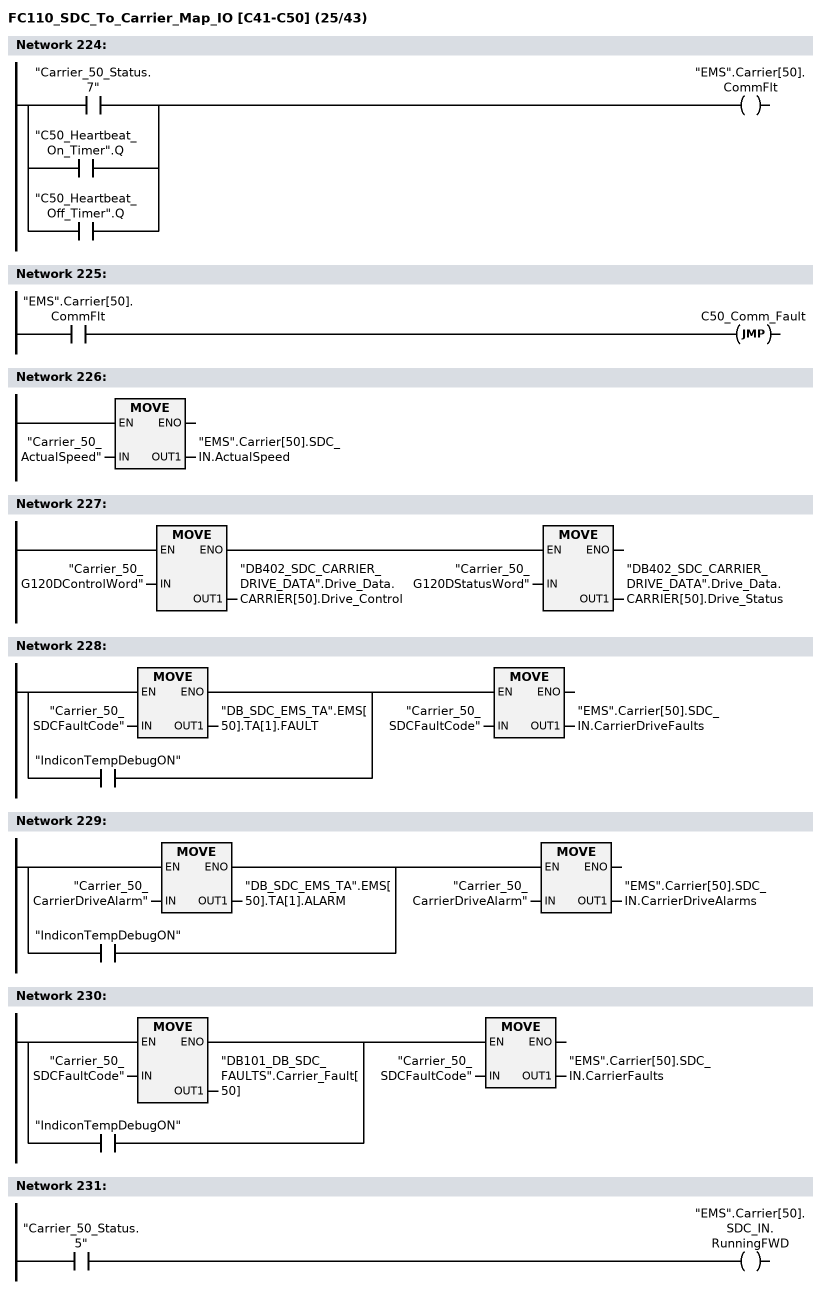
   RUNG wire#powerrail
      Contact( "Carrier_50_Status.7" )
      wire#w1
      Coil( "EMS".Carrier[50].CommFlt )
   END_RUNG
   RUNG wire#powerrail
      Contact( "C50_Heartbeat_On_Timer".Q )
   END_RUNG wire#w1
   RUNG wire#powerrail
      Contact( "C50_Heartbeat_Off_Timer".Q )
   END_RUNG wire#w1
   // the same network as SCL:
   "EMS".Carrier[50].CommFlt := "Carrier_50_Status.7" OR "C50_Heartbeat_On_Timer".Q OR "C50_Heartbeat_Off_Timer".Q;
END_REGION

REGION Network 225
   RUNG wire#powerrail
      Contact( "EMS".Carrier[50].CommFlt )
      JumpCoil( C50_Comm_Fault )
   END_RUNG
   // the same network as SCL:
   IF "EMS".Carrier[50].CommFlt THEN GOTO C50_Comm_Fault; END_IF;
END_REGION

REGION Network 226
   RUNG wire#powerrail
      Move(in := "Carrier_50_ActualSpeed", out1 => "EMS".Carrier[50].SDC_IN.ActualSpeed)
   END_RUNG
   // the same network as SCL:
   "EMS".Carrier[50].SDC_IN.ActualSpeed := "Carrier_50_ActualSpeed";
END_REGION

REGION Network 227
   RUNG wire#powerrail
      Move(in := "Carrier_50_G120DControlWord", out1 => "DB402_SDC_CARRIER_DRIVE_DATA".Drive_Data.CARRIER[50].Drive_Control)
      Move(in := "Carrier_50_G120DStatusWord", out1 => "DB402_SDC_CARRIER_DRIVE_DATA".Drive_Data.CARRIER[50].Drive_Status)
   END_RUNG
   // the same network as SCL:
   "DB402_SDC_CARRIER_DRIVE_DATA".Drive_Data.CARRIER[50].Drive_Control := "Carrier_50_G120DControlWord";
   "DB402_SDC_CARRIER_DRIVE_DATA".Drive_Data.CARRIER[50].Drive_Status := "Carrier_50_G120DStatusWord";
END_REGION

REGION Network 228
   RUNG wire#powerrail
      Move(in := "Carrier_50_SDCFaultCode", out1 => "DB_SDC_EMS_TA".EMS[50].TA[1].FAULT)
      wire#w1
      Move(in := "Carrier_50_SDCFaultCode", out1 => "EMS".Carrier[50].SDC_IN.CarrierDriveFaults)
   END_RUNG
   RUNG wire#powerrail
      Contact( "IndiconTempDebugON" )
   END_RUNG wire#w1
   // the same network as SCL:
   "DB_SDC_EMS_TA".EMS[50].TA[1].FAULT := "Carrier_50_SDCFaultCode";
   IF TRUE OR "IndiconTempDebugON" THEN
       "EMS".Carrier[50].SDC_IN.CarrierDriveFaults := "Carrier_50_SDCFaultCode";
   END_IF;
END_REGION

REGION Network 229
   RUNG wire#powerrail
      Move(in := "Carrier_50_CarrierDriveAlarm", out1 => "DB_SDC_EMS_TA".EMS[50].TA[1].ALARM)
      wire#w1
      Move(in := "Carrier_50_CarrierDriveAlarm", out1 => "EMS".Carrier[50].SDC_IN.CarrierDriveAlarms)
   END_RUNG
   RUNG wire#powerrail
      Contact( "IndiconTempDebugON" )
   END_RUNG wire#w1
   // the same network as SCL:
   "DB_SDC_EMS_TA".EMS[50].TA[1].ALARM := "Carrier_50_CarrierDriveAlarm";
   IF TRUE OR "IndiconTempDebugON" THEN
       "EMS".Carrier[50].SDC_IN.CarrierDriveAlarms := "Carrier_50_CarrierDriveAlarm";
   END_IF;
END_REGION

REGION Network 230
   RUNG wire#powerrail
      Move(in := "Carrier_50_SDCFaultCode", out1 => "DB101_DB_SDC_FAULTS".Carrier_Fault[50])
      wire#w1
      Move(in := "Carrier_50_SDCFaultCode", out1 => "EMS".Carrier[50].SDC_IN.CarrierFaults)
   END_RUNG
   RUNG wire#powerrail
      Contact( "IndiconTempDebugON" )
   END_RUNG wire#w1
   // the same network as SCL:
   "DB101_DB_SDC_FAULTS".Carrier_Fault[50] := "Carrier_50_SDCFaultCode";
   IF TRUE OR "IndiconTempDebugON" THEN
       "EMS".Carrier[50].SDC_IN.CarrierFaults := "Carrier_50_SDCFaultCode";
   END_IF;
END_REGION

REGION Network 231
   RUNG wire#powerrail
      Contact( "Carrier_50_Status.5" )
      Coil( "EMS".Carrier[50].SDC_IN.RunningFWD )
   END_RUNG
   // the same network as SCL:
   "EMS".Carrier[50].SDC_IN.RunningFWD := "Carrier_50_Status.5";
END_REGION

REGION Network 232
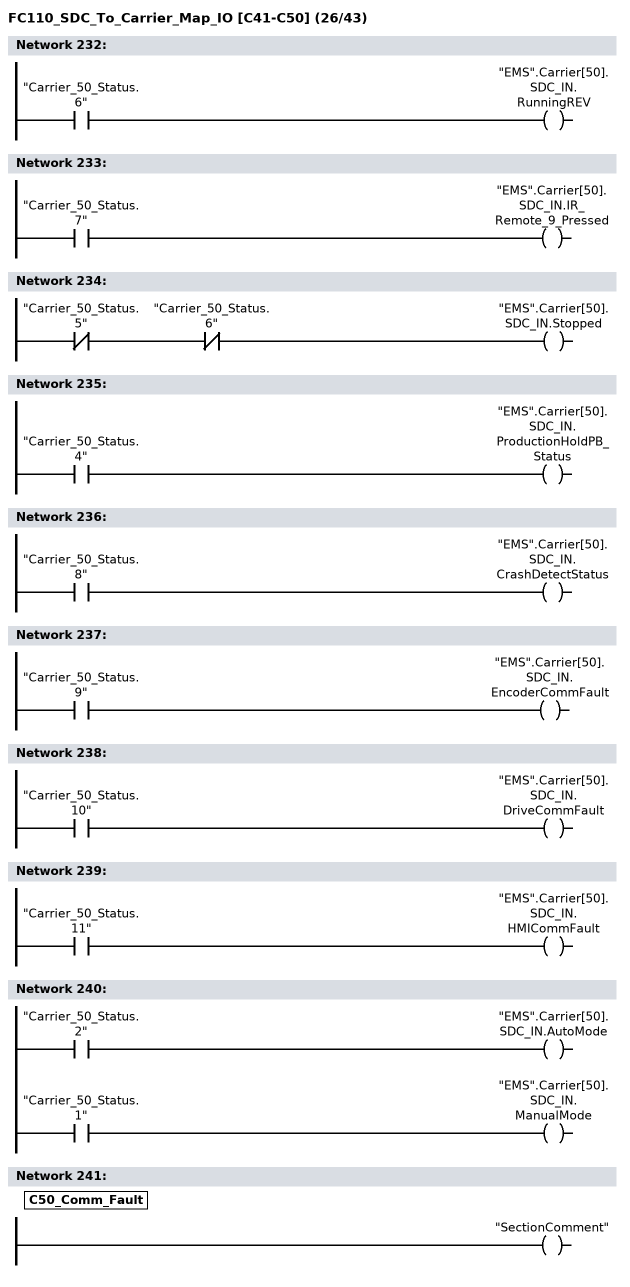
   RUNG wire#powerrail
      Contact( "Carrier_50_Status.6" )
      Coil( "EMS".Carrier[50].SDC_IN.RunningREV )
   END_RUNG
   // the same network as SCL:
   "EMS".Carrier[50].SDC_IN.RunningREV := "Carrier_50_Status.6";
END_REGION

REGION Network 233
   RUNG wire#powerrail
      Contact( "Carrier_50_Status.7" )
      Coil( "EMS".Carrier[50].SDC_IN.IR_Remote_9_Pressed )
   END_RUNG
   // the same network as SCL:
   "EMS".Carrier[50].SDC_IN.IR_Remote_9_Pressed := "Carrier_50_Status.7";
END_REGION

REGION Network 234
   RUNG wire#powerrail
      I_Contact( "Carrier_50_Status.5" )
      I_Contact( "Carrier_50_Status.6" )
      Coil( "EMS".Carrier[50].SDC_IN.Stopped )
   END_RUNG
   // the same network as SCL:
   "EMS".Carrier[50].SDC_IN.Stopped := NOT "Carrier_50_Status.5" AND NOT "Carrier_50_Status.6";
END_REGION

REGION Network 235
   RUNG wire#powerrail
      Contact( "Carrier_50_Status.4" )
      Coil( "EMS".Carrier[50].SDC_IN.ProductionHoldPB_Status )
   END_RUNG
   // the same network as SCL:
   "EMS".Carrier[50].SDC_IN.ProductionHoldPB_Status := "Carrier_50_Status.4";
END_REGION

REGION Network 236
   RUNG wire#powerrail
      Contact( "Carrier_50_Status.8" )
      Coil( "EMS".Carrier[50].SDC_IN.CrashDetectStatus )
   END_RUNG
   // the same network as SCL:
   "EMS".Carrier[50].SDC_IN.CrashDetectStatus := "Carrier_50_Status.8";
END_REGION

REGION Network 237
   RUNG wire#powerrail
      Contact( "Carrier_50_Status.9" )
      Coil( "EMS".Carrier[50].SDC_IN.EncoderCommFault )
   END_RUNG
   // the same network as SCL:
   "EMS".Carrier[50].SDC_IN.EncoderCommFault := "Carrier_50_Status.9";
END_REGION

REGION Network 238
   RUNG wire#powerrail
      Contact( "Carrier_50_Status.10" )
      Coil( "EMS".Carrier[50].SDC_IN.DriveCommFault )
   END_RUNG
   // the same network as SCL:
   "EMS".Carrier[50].SDC_IN.DriveCommFault := "Carrier_50_Status.10";
END_REGION

REGION Network 239
   RUNG wire#powerrail
      Contact( "Carrier_50_Status.11" )
      Coil( "EMS".Carrier[50].SDC_IN.HMICommFault )
   END_RUNG
   // the same network as SCL:
   "EMS".Carrier[50].SDC_IN.HMICommFault := "Carrier_50_Status.11";
END_REGION

REGION Network 240
   RUNG wire#powerrail
      Contact( "Carrier_50_Status.2" )
      Coil( "EMS".Carrier[50].SDC_IN.AutoMode )
   END_RUNG
   RUNG wire#powerrail
      Contact( "Carrier_50_Status.1" )
      Coil( "EMS".Carrier[50].SDC_IN.ManualMode )
   END_RUNG
   // the same network as SCL:
   "EMS".Carrier[50].SDC_IN.AutoMode := "Carrier_50_Status.2";
   "EMS".Carrier[50].SDC_IN.ManualMode := "Carrier_50_Status.1";
END_REGION

REGION Network 241
   Label( C50_Comm_Fault )
   RUNG wire#powerrail
      Coil( "SectionComment" )
   END_RUNG
   // the same network as SCL:
   C50_Comm_Fault:
   "SectionComment" := TRUE;
END_REGION

REGION Network 242
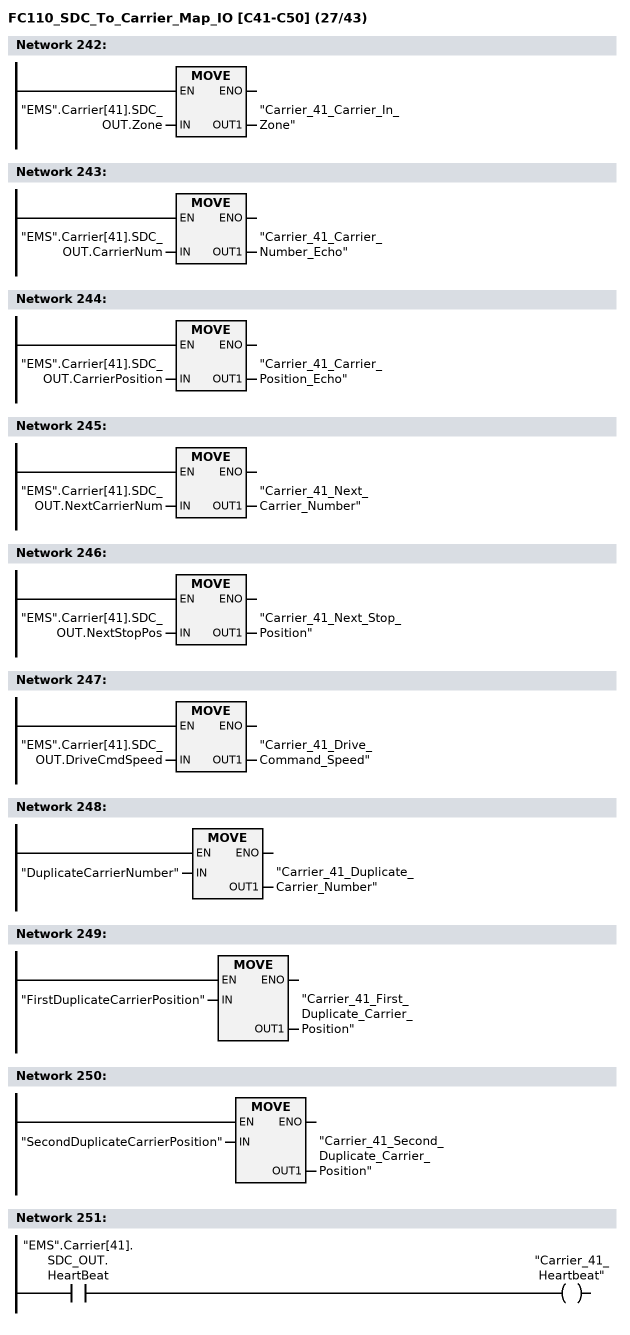
   RUNG wire#powerrail
      Move(in := "EMS".Carrier[41].SDC_OUT.Zone, out1 => "Carrier_41_Carrier_In_Zone")
   END_RUNG
   // the same network as SCL:
   "Carrier_41_Carrier_In_Zone" := "EMS".Carrier[41].SDC_OUT.Zone;
END_REGION

REGION Network 243
   RUNG wire#powerrail
      Move(in := "EMS".Carrier[41].SDC_OUT.CarrierNum, out1 => "Carrier_41_Carrier_Number_Echo")
   END_RUNG
   // the same network as SCL:
   "Carrier_41_Carrier_Number_Echo" := "EMS".Carrier[41].SDC_OUT.CarrierNum;
END_REGION

REGION Network 244
   RUNG wire#powerrail
      Move(in := "EMS".Carrier[41].SDC_OUT.CarrierPosition, out1 => "Carrier_41_Carrier_Position_Echo")
   END_RUNG
   // the same network as SCL:
   "Carrier_41_Carrier_Position_Echo" := "EMS".Carrier[41].SDC_OUT.CarrierPosition;
END_REGION

REGION Network 245
   RUNG wire#powerrail
      Move(in := "EMS".Carrier[41].SDC_OUT.NextCarrierNum, out1 => "Carrier_41_Next_Carrier_Number")
   END_RUNG
   // the same network as SCL:
   "Carrier_41_Next_Carrier_Number" := "EMS".Carrier[41].SDC_OUT.NextCarrierNum;
END_REGION

REGION Network 246
   RUNG wire#powerrail
      Move(in := "EMS".Carrier[41].SDC_OUT.NextStopPos, out1 => "Carrier_41_Next_Stop_Position")
   END_RUNG
   // the same network as SCL:
   "Carrier_41_Next_Stop_Position" := "EMS".Carrier[41].SDC_OUT.NextStopPos;
END_REGION

REGION Network 247
   RUNG wire#powerrail
      Move(in := "EMS".Carrier[41].SDC_OUT.DriveCmdSpeed, out1 => "Carrier_41_Drive_Command_Speed")
   END_RUNG
   // the same network as SCL:
   "Carrier_41_Drive_Command_Speed" := "EMS".Carrier[41].SDC_OUT.DriveCmdSpeed;
END_REGION

REGION Network 248
   RUNG wire#powerrail
      Move(in := "DuplicateCarrierNumber", out1 => "Carrier_41_Duplicate_Carrier_Number")
   END_RUNG
   // the same network as SCL:
   "Carrier_41_Duplicate_Carrier_Number" := "DuplicateCarrierNumber";
END_REGION

REGION Network 249
   RUNG wire#powerrail
      Move(in := "FirstDuplicateCarrierPosition", out1 => "Carrier_41_First_Duplicate_Carrier_Position")
   END_RUNG
   // the same network as SCL:
   "Carrier_41_First_Duplicate_Carrier_Position" := "FirstDuplicateCarrierPosition";
END_REGION

REGION Network 250
   RUNG wire#powerrail
      Move(in := "SecondDuplicateCarrierPosition", out1 => "Carrier_41_Second_Duplicate_Carrier_Position")
   END_RUNG
   // the same network as SCL:
   "Carrier_41_Second_Duplicate_Carrier_Position" := "SecondDuplicateCarrierPosition";
END_REGION

REGION Network 251
   RUNG wire#powerrail
      Contact( "EMS".Carrier[41].SDC_OUT.HeartBeat )
      Coil( "Carrier_41_Heartbeat" )
   END_RUNG
   // the same network as SCL:
   "Carrier_41_Heartbeat" := "EMS".Carrier[41].SDC_OUT.HeartBeat;
END_REGION

REGION Network 252
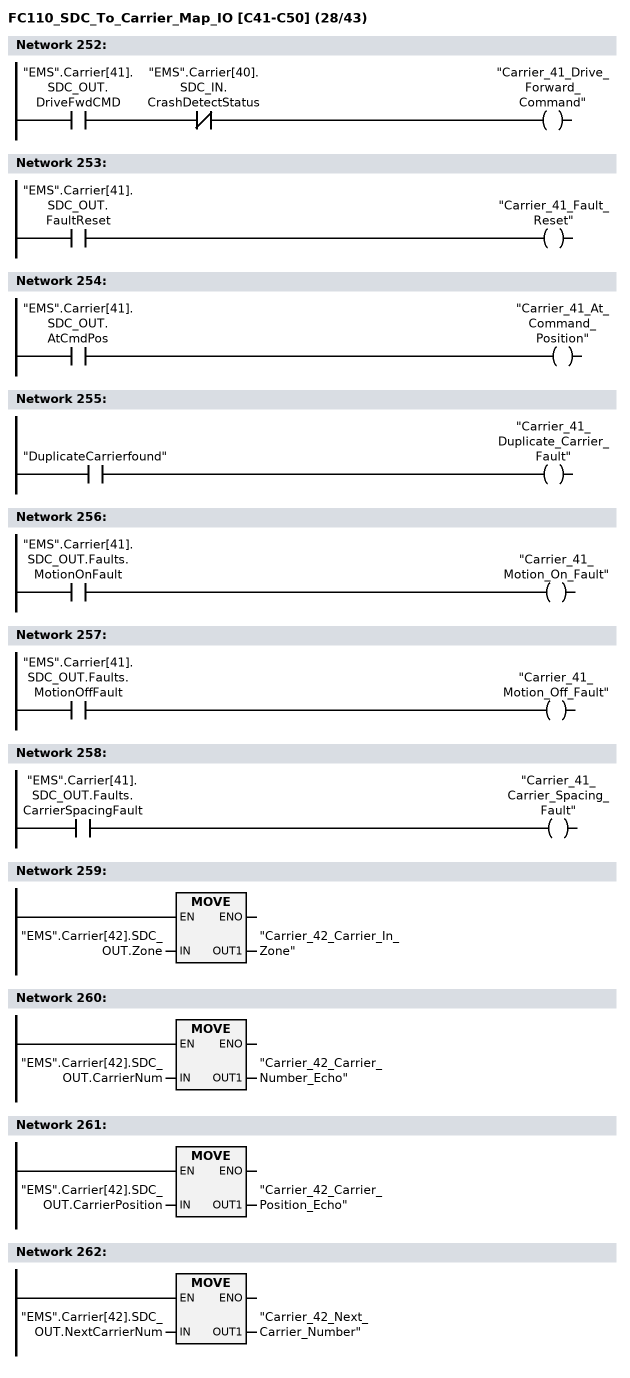
   RUNG wire#powerrail
      Contact( "EMS".Carrier[41].SDC_OUT.DriveFwdCMD )
      I_Contact( "EMS".Carrier[40].SDC_IN.CrashDetectStatus )
      Coil( "Carrier_41_Drive_Forward_Command" )
   END_RUNG
   // the same network as SCL:
   "Carrier_41_Drive_Forward_Command" := "EMS".Carrier[41].SDC_OUT.DriveFwdCMD AND NOT "EMS".Carrier[40].SDC_IN.CrashDetectStatus;
END_REGION

REGION Network 253
   RUNG wire#powerrail
      Contact( "EMS".Carrier[41].SDC_OUT.FaultReset )
      Coil( "Carrier_41_Fault_Reset" )
   END_RUNG
   // the same network as SCL:
   "Carrier_41_Fault_Reset" := "EMS".Carrier[41].SDC_OUT.FaultReset;
END_REGION

REGION Network 254
   RUNG wire#powerrail
      Contact( "EMS".Carrier[41].SDC_OUT.AtCmdPos )
      Coil( "Carrier_41_At_Command_Position" )
   END_RUNG
   // the same network as SCL:
   "Carrier_41_At_Command_Position" := "EMS".Carrier[41].SDC_OUT.AtCmdPos;
END_REGION

REGION Network 255
   RUNG wire#powerrail
      Contact( "DuplicateCarrierfound" )
      Coil( "Carrier_41_Duplicate_Carrier_Fault" )
   END_RUNG
   // the same network as SCL:
   "Carrier_41_Duplicate_Carrier_Fault" := "DuplicateCarrierfound";
END_REGION

REGION Network 256
   RUNG wire#powerrail
      Contact( "EMS".Carrier[41].SDC_OUT.Faults.MotionOnFault )
      Coil( "Carrier_41_Motion_On_Fault" )
   END_RUNG
   // the same network as SCL:
   "Carrier_41_Motion_On_Fault" := "EMS".Carrier[41].SDC_OUT.Faults.MotionOnFault;
END_REGION

REGION Network 257
   RUNG wire#powerrail
      Contact( "EMS".Carrier[41].SDC_OUT.Faults.MotionOffFault )
      Coil( "Carrier_41_Motion_Off_Fault" )
   END_RUNG
   // the same network as SCL:
   "Carrier_41_Motion_Off_Fault" := "EMS".Carrier[41].SDC_OUT.Faults.MotionOffFault;
END_REGION

REGION Network 258
   RUNG wire#powerrail
      Contact( "EMS".Carrier[41].SDC_OUT.Faults.CarrierSpacingFault )
      Coil( "Carrier_41_Carrier_Spacing_Fault" )
   END_RUNG
   // the same network as SCL:
   "Carrier_41_Carrier_Spacing_Fault" := "EMS".Carrier[41].SDC_OUT.Faults.CarrierSpacingFault;
END_REGION

REGION Network 259
   RUNG wire#powerrail
      Move(in := "EMS".Carrier[42].SDC_OUT.Zone, out1 => "Carrier_42_Carrier_In_Zone")
   END_RUNG
   // the same network as SCL:
   "Carrier_42_Carrier_In_Zone" := "EMS".Carrier[42].SDC_OUT.Zone;
END_REGION

REGION Network 260
   RUNG wire#powerrail
      Move(in := "EMS".Carrier[42].SDC_OUT.CarrierNum, out1 => "Carrier_42_Carrier_Number_Echo")
   END_RUNG
   // the same network as SCL:
   "Carrier_42_Carrier_Number_Echo" := "EMS".Carrier[42].SDC_OUT.CarrierNum;
END_REGION

REGION Network 261
   RUNG wire#powerrail
      Move(in := "EMS".Carrier[42].SDC_OUT.CarrierPosition, out1 => "Carrier_42_Carrier_Position_Echo")
   END_RUNG
   // the same network as SCL:
   "Carrier_42_Carrier_Position_Echo" := "EMS".Carrier[42].SDC_OUT.CarrierPosition;
END_REGION

REGION Network 262
   RUNG wire#powerrail
      Move(in := "EMS".Carrier[42].SDC_OUT.NextCarrierNum, out1 => "Carrier_42_Next_Carrier_Number")
   END_RUNG
   // the same network as SCL:
   "Carrier_42_Next_Carrier_Number" := "EMS".Carrier[42].SDC_OUT.NextCarrierNum;
END_REGION

REGION Network 263
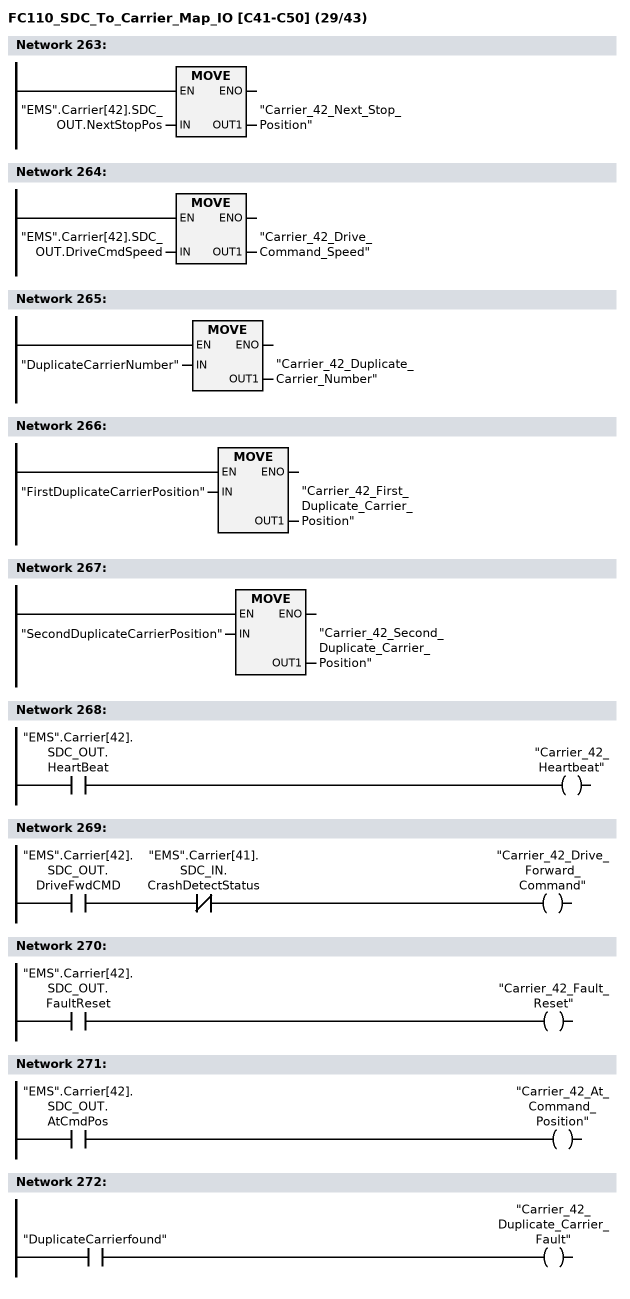
   RUNG wire#powerrail
      Move(in := "EMS".Carrier[42].SDC_OUT.NextStopPos, out1 => "Carrier_42_Next_Stop_Position")
   END_RUNG
   // the same network as SCL:
   "Carrier_42_Next_Stop_Position" := "EMS".Carrier[42].SDC_OUT.NextStopPos;
END_REGION

REGION Network 264
   RUNG wire#powerrail
      Move(in := "EMS".Carrier[42].SDC_OUT.DriveCmdSpeed, out1 => "Carrier_42_Drive_Command_Speed")
   END_RUNG
   // the same network as SCL:
   "Carrier_42_Drive_Command_Speed" := "EMS".Carrier[42].SDC_OUT.DriveCmdSpeed;
END_REGION

REGION Network 265
   RUNG wire#powerrail
      Move(in := "DuplicateCarrierNumber", out1 => "Carrier_42_Duplicate_Carrier_Number")
   END_RUNG
   // the same network as SCL:
   "Carrier_42_Duplicate_Carrier_Number" := "DuplicateCarrierNumber";
END_REGION

REGION Network 266
   RUNG wire#powerrail
      Move(in := "FirstDuplicateCarrierPosition", out1 => "Carrier_42_First_Duplicate_Carrier_Position")
   END_RUNG
   // the same network as SCL:
   "Carrier_42_First_Duplicate_Carrier_Position" := "FirstDuplicateCarrierPosition";
END_REGION

REGION Network 267
   RUNG wire#powerrail
      Move(in := "SecondDuplicateCarrierPosition", out1 => "Carrier_42_Second_Duplicate_Carrier_Position")
   END_RUNG
   // the same network as SCL:
   "Carrier_42_Second_Duplicate_Carrier_Position" := "SecondDuplicateCarrierPosition";
END_REGION

REGION Network 268
   RUNG wire#powerrail
      Contact( "EMS".Carrier[42].SDC_OUT.HeartBeat )
      Coil( "Carrier_42_Heartbeat" )
   END_RUNG
   // the same network as SCL:
   "Carrier_42_Heartbeat" := "EMS".Carrier[42].SDC_OUT.HeartBeat;
END_REGION

REGION Network 269
   RUNG wire#powerrail
      Contact( "EMS".Carrier[42].SDC_OUT.DriveFwdCMD )
      I_Contact( "EMS".Carrier[41].SDC_IN.CrashDetectStatus )
      Coil( "Carrier_42_Drive_Forward_Command" )
   END_RUNG
   // the same network as SCL:
   "Carrier_42_Drive_Forward_Command" := "EMS".Carrier[42].SDC_OUT.DriveFwdCMD AND NOT "EMS".Carrier[41].SDC_IN.CrashDetectStatus;
END_REGION

REGION Network 270
   RUNG wire#powerrail
      Contact( "EMS".Carrier[42].SDC_OUT.FaultReset )
      Coil( "Carrier_42_Fault_Reset" )
   END_RUNG
   // the same network as SCL:
   "Carrier_42_Fault_Reset" := "EMS".Carrier[42].SDC_OUT.FaultReset;
END_REGION

REGION Network 271
   RUNG wire#powerrail
      Contact( "EMS".Carrier[42].SDC_OUT.AtCmdPos )
      Coil( "Carrier_42_At_Command_Position" )
   END_RUNG
   // the same network as SCL:
   "Carrier_42_At_Command_Position" := "EMS".Carrier[42].SDC_OUT.AtCmdPos;
END_REGION

REGION Network 272
   RUNG wire#powerrail
      Contact( "DuplicateCarrierfound" )
      Coil( "Carrier_42_Duplicate_Carrier_Fault" )
   END_RUNG
   // the same network as SCL:
   "Carrier_42_Duplicate_Carrier_Fault" := "DuplicateCarrierfound";
END_REGION

REGION Network 273
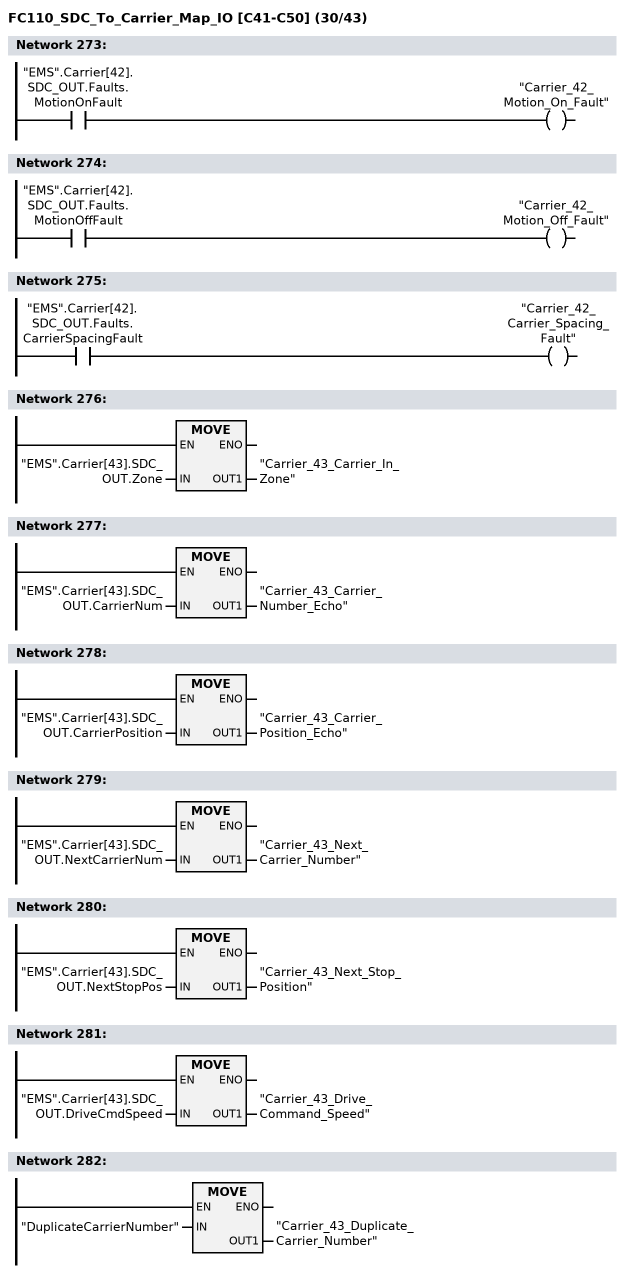
   RUNG wire#powerrail
      Contact( "EMS".Carrier[42].SDC_OUT.Faults.MotionOnFault )
      Coil( "Carrier_42_Motion_On_Fault" )
   END_RUNG
   // the same network as SCL:
   "Carrier_42_Motion_On_Fault" := "EMS".Carrier[42].SDC_OUT.Faults.MotionOnFault;
END_REGION

REGION Network 274
   RUNG wire#powerrail
      Contact( "EMS".Carrier[42].SDC_OUT.Faults.MotionOffFault )
      Coil( "Carrier_42_Motion_Off_Fault" )
   END_RUNG
   // the same network as SCL:
   "Carrier_42_Motion_Off_Fault" := "EMS".Carrier[42].SDC_OUT.Faults.MotionOffFault;
END_REGION

REGION Network 275
   RUNG wire#powerrail
      Contact( "EMS".Carrier[42].SDC_OUT.Faults.CarrierSpacingFault )
      Coil( "Carrier_42_Carrier_Spacing_Fault" )
   END_RUNG
   // the same network as SCL:
   "Carrier_42_Carrier_Spacing_Fault" := "EMS".Carrier[42].SDC_OUT.Faults.CarrierSpacingFault;
END_REGION

REGION Network 276
   RUNG wire#powerrail
      Move(in := "EMS".Carrier[43].SDC_OUT.Zone, out1 => "Carrier_43_Carrier_In_Zone")
   END_RUNG
   // the same network as SCL:
   "Carrier_43_Carrier_In_Zone" := "EMS".Carrier[43].SDC_OUT.Zone;
END_REGION

REGION Network 277
   RUNG wire#powerrail
      Move(in := "EMS".Carrier[43].SDC_OUT.CarrierNum, out1 => "Carrier_43_Carrier_Number_Echo")
   END_RUNG
   // the same network as SCL:
   "Carrier_43_Carrier_Number_Echo" := "EMS".Carrier[43].SDC_OUT.CarrierNum;
END_REGION

REGION Network 278
   RUNG wire#powerrail
      Move(in := "EMS".Carrier[43].SDC_OUT.CarrierPosition, out1 => "Carrier_43_Carrier_Position_Echo")
   END_RUNG
   // the same network as SCL:
   "Carrier_43_Carrier_Position_Echo" := "EMS".Carrier[43].SDC_OUT.CarrierPosition;
END_REGION

REGION Network 279
   RUNG wire#powerrail
      Move(in := "EMS".Carrier[43].SDC_OUT.NextCarrierNum, out1 => "Carrier_43_Next_Carrier_Number")
   END_RUNG
   // the same network as SCL:
   "Carrier_43_Next_Carrier_Number" := "EMS".Carrier[43].SDC_OUT.NextCarrierNum;
END_REGION

REGION Network 280
   RUNG wire#powerrail
      Move(in := "EMS".Carrier[43].SDC_OUT.NextStopPos, out1 => "Carrier_43_Next_Stop_Position")
   END_RUNG
   // the same network as SCL:
   "Carrier_43_Next_Stop_Position" := "EMS".Carrier[43].SDC_OUT.NextStopPos;
END_REGION

REGION Network 281
   RUNG wire#powerrail
      Move(in := "EMS".Carrier[43].SDC_OUT.DriveCmdSpeed, out1 => "Carrier_43_Drive_Command_Speed")
   END_RUNG
   // the same network as SCL:
   "Carrier_43_Drive_Command_Speed" := "EMS".Carrier[43].SDC_OUT.DriveCmdSpeed;
END_REGION

REGION Network 282
   RUNG wire#powerrail
      Move(in := "DuplicateCarrierNumber", out1 => "Carrier_43_Duplicate_Carrier_Number")
   END_RUNG
   // the same network as SCL:
   "Carrier_43_Duplicate_Carrier_Number" := "DuplicateCarrierNumber";
END_REGION

REGION Network 283
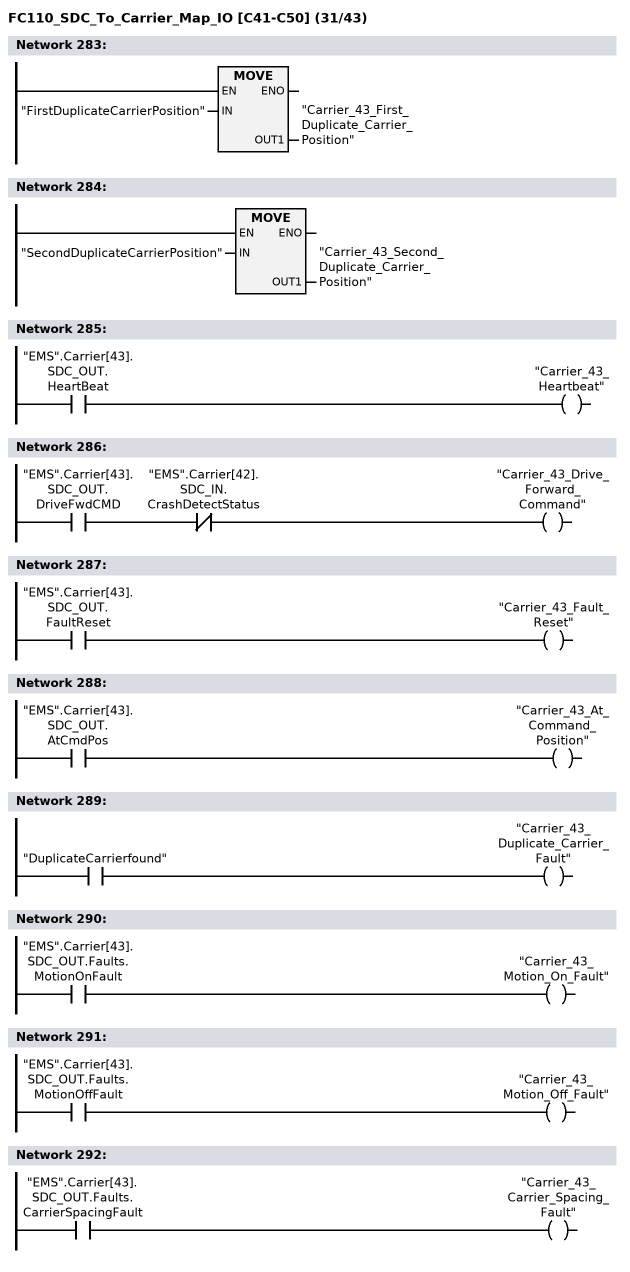
   RUNG wire#powerrail
      Move(in := "FirstDuplicateCarrierPosition", out1 => "Carrier_43_First_Duplicate_Carrier_Position")
   END_RUNG
   // the same network as SCL:
   "Carrier_43_First_Duplicate_Carrier_Position" := "FirstDuplicateCarrierPosition";
END_REGION

REGION Network 284
   RUNG wire#powerrail
      Move(in := "SecondDuplicateCarrierPosition", out1 => "Carrier_43_Second_Duplicate_Carrier_Position")
   END_RUNG
   // the same network as SCL:
   "Carrier_43_Second_Duplicate_Carrier_Position" := "SecondDuplicateCarrierPosition";
END_REGION

REGION Network 285
   RUNG wire#powerrail
      Contact( "EMS".Carrier[43].SDC_OUT.HeartBeat )
      Coil( "Carrier_43_Heartbeat" )
   END_RUNG
   // the same network as SCL:
   "Carrier_43_Heartbeat" := "EMS".Carrier[43].SDC_OUT.HeartBeat;
END_REGION

REGION Network 286
   RUNG wire#powerrail
      Contact( "EMS".Carrier[43].SDC_OUT.DriveFwdCMD )
      I_Contact( "EMS".Carrier[42].SDC_IN.CrashDetectStatus )
      Coil( "Carrier_43_Drive_Forward_Command" )
   END_RUNG
   // the same network as SCL:
   "Carrier_43_Drive_Forward_Command" := "EMS".Carrier[43].SDC_OUT.DriveFwdCMD AND NOT "EMS".Carrier[42].SDC_IN.CrashDetectStatus;
END_REGION

REGION Network 287
   RUNG wire#powerrail
      Contact( "EMS".Carrier[43].SDC_OUT.FaultReset )
      Coil( "Carrier_43_Fault_Reset" )
   END_RUNG
   // the same network as SCL:
   "Carrier_43_Fault_Reset" := "EMS".Carrier[43].SDC_OUT.FaultReset;
END_REGION

REGION Network 288
   RUNG wire#powerrail
      Contact( "EMS".Carrier[43].SDC_OUT.AtCmdPos )
      Coil( "Carrier_43_At_Command_Position" )
   END_RUNG
   // the same network as SCL:
   "Carrier_43_At_Command_Position" := "EMS".Carrier[43].SDC_OUT.AtCmdPos;
END_REGION

REGION Network 289
   RUNG wire#powerrail
      Contact( "DuplicateCarrierfound" )
      Coil( "Carrier_43_Duplicate_Carrier_Fault" )
   END_RUNG
   // the same network as SCL:
   "Carrier_43_Duplicate_Carrier_Fault" := "DuplicateCarrierfound";
END_REGION

REGION Network 290
   RUNG wire#powerrail
      Contact( "EMS".Carrier[43].SDC_OUT.Faults.MotionOnFault )
      Coil( "Carrier_43_Motion_On_Fault" )
   END_RUNG
   // the same network as SCL:
   "Carrier_43_Motion_On_Fault" := "EMS".Carrier[43].SDC_OUT.Faults.MotionOnFault;
END_REGION

REGION Network 291
   RUNG wire#powerrail
      Contact( "EMS".Carrier[43].SDC_OUT.Faults.MotionOffFault )
      Coil( "Carrier_43_Motion_Off_Fault" )
   END_RUNG
   // the same network as SCL:
   "Carrier_43_Motion_Off_Fault" := "EMS".Carrier[43].SDC_OUT.Faults.MotionOffFault;
END_REGION

REGION Network 292
   RUNG wire#powerrail
      Contact( "EMS".Carrier[43].SDC_OUT.Faults.CarrierSpacingFault )
      Coil( "Carrier_43_Carrier_Spacing_Fault" )
   END_RUNG
   // the same network as SCL:
   "Carrier_43_Carrier_Spacing_Fault" := "EMS".Carrier[43].SDC_OUT.Faults.CarrierSpacingFault;
END_REGION

REGION Network 293
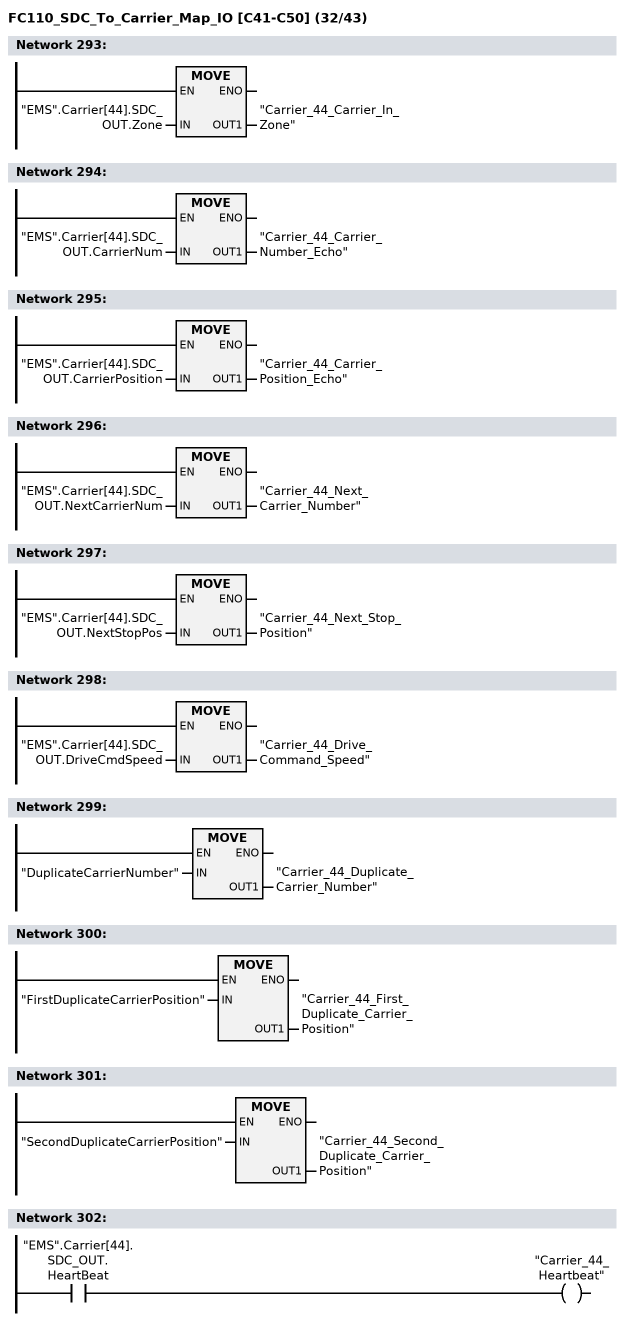
   RUNG wire#powerrail
      Move(in := "EMS".Carrier[44].SDC_OUT.Zone, out1 => "Carrier_44_Carrier_In_Zone")
   END_RUNG
   // the same network as SCL:
   "Carrier_44_Carrier_In_Zone" := "EMS".Carrier[44].SDC_OUT.Zone;
END_REGION

REGION Network 294
   RUNG wire#powerrail
      Move(in := "EMS".Carrier[44].SDC_OUT.CarrierNum, out1 => "Carrier_44_Carrier_Number_Echo")
   END_RUNG
   // the same network as SCL:
   "Carrier_44_Carrier_Number_Echo" := "EMS".Carrier[44].SDC_OUT.CarrierNum;
END_REGION

REGION Network 295
   RUNG wire#powerrail
      Move(in := "EMS".Carrier[44].SDC_OUT.CarrierPosition, out1 => "Carrier_44_Carrier_Position_Echo")
   END_RUNG
   // the same network as SCL:
   "Carrier_44_Carrier_Position_Echo" := "EMS".Carrier[44].SDC_OUT.CarrierPosition;
END_REGION

REGION Network 296
   RUNG wire#powerrail
      Move(in := "EMS".Carrier[44].SDC_OUT.NextCarrierNum, out1 => "Carrier_44_Next_Carrier_Number")
   END_RUNG
   // the same network as SCL:
   "Carrier_44_Next_Carrier_Number" := "EMS".Carrier[44].SDC_OUT.NextCarrierNum;
END_REGION

REGION Network 297
   RUNG wire#powerrail
      Move(in := "EMS".Carrier[44].SDC_OUT.NextStopPos, out1 => "Carrier_44_Next_Stop_Position")
   END_RUNG
   // the same network as SCL:
   "Carrier_44_Next_Stop_Position" := "EMS".Carrier[44].SDC_OUT.NextStopPos;
END_REGION

REGION Network 298
   RUNG wire#powerrail
      Move(in := "EMS".Carrier[44].SDC_OUT.DriveCmdSpeed, out1 => "Carrier_44_Drive_Command_Speed")
   END_RUNG
   // the same network as SCL:
   "Carrier_44_Drive_Command_Speed" := "EMS".Carrier[44].SDC_OUT.DriveCmdSpeed;
END_REGION

REGION Network 299
   RUNG wire#powerrail
      Move(in := "DuplicateCarrierNumber", out1 => "Carrier_44_Duplicate_Carrier_Number")
   END_RUNG
   // the same network as SCL:
   "Carrier_44_Duplicate_Carrier_Number" := "DuplicateCarrierNumber";
END_REGION

REGION Network 300
   RUNG wire#powerrail
      Move(in := "FirstDuplicateCarrierPosition", out1 => "Carrier_44_First_Duplicate_Carrier_Position")
   END_RUNG
   // the same network as SCL:
   "Carrier_44_First_Duplicate_Carrier_Position" := "FirstDuplicateCarrierPosition";
END_REGION

REGION Network 301
   RUNG wire#powerrail
      Move(in := "SecondDuplicateCarrierPosition", out1 => "Carrier_44_Second_Duplicate_Carrier_Position")
   END_RUNG
   // the same network as SCL:
   "Carrier_44_Second_Duplicate_Carrier_Position" := "SecondDuplicateCarrierPosition";
END_REGION

REGION Network 302
   RUNG wire#powerrail
      Contact( "EMS".Carrier[44].SDC_OUT.HeartBeat )
      Coil( "Carrier_44_Heartbeat" )
   END_RUNG
   // the same network as SCL:
   "Carrier_44_Heartbeat" := "EMS".Carrier[44].SDC_OUT.HeartBeat;
END_REGION

REGION Network 303